(* Logix 5000 project; controller FV vendor 1 type 14 code 217 rev 31.11; software revision 31.00; part 51 of 63 *)
(* tags used below, declared in another part *)
   CWD : CHECKWORD_FLAGS;
   FV_AV1 : PlantItem;   // AV1
   FV_B32 : INT[255];   // PITCH_FLGS YSV pitching control flags
   FV_B32_0_2_OutputBit : BOOL;
   fv_data_file_value_to_move : DINT;
   FV_N12 : INT[255];   // SYS_PARMS System Parameter Fil e
   FV_N141 : INT[255];   // YSV1 DATA
   FV_N142 : INT[255];   // YSV2 DATA
   FV_N143 : INT[255];   // YSV3 DATA
   FV_N30 : INT[255];   // PITCH<PC YSV Pitching data fr om PC
   FV_N31 : INT[255];   // PITCH>PC YSV Pitching data at o PC and control reg isters
   FV_N34 : INT[255];   // PITCH_SV YSV pitching data sa ve file to PC
   FV_N50 : INT[255];   // WASTE<PC
   FV_T33 : TIMER[10];
   FV_YSV1_WTX01_AI : PlantItem;   // YSV1_WTX01
   FV_YSV2_WTX01_AI : PlantItem;   // YSV2_WTX01
   FV_YSV2O : PlantItem;   // YSV2O
   FV_YSV3_WTX01_AI : PlantItem;   // YSV3_WTX01
   FV_YSV3O : PlantItem;   // YSV3O
   FV_YSVPitching_AmountAtEnd : REAL;
   Pitching_transaction_log_delay : DINT;
(* FV_Common, continued *)

ROUTINE FV_PITCH_CP_16   (* ladder *)
   // Reset command interpreter step counter
   0: XIC(S:FS)CLR(FV_N31[16]);
   // RESET
   1: EQU(FV_N31[16],0)MCR();
   2: OTU(FV_B32[0].0);
   3: OTU(FV_B32[0].1);
   4: OTU(FV_B32[0].8);
   5: FLL(0,FV_N31[0],16);
   // Set PCparameter buffer to 'Null' value
   6: FLL(-32768,FV_N30[1],7);
   7: CLR(FV_N30[0]);
   8: MOV(1,FV_N31[16]);
   9: MCR();
   // ALLOW STARTUP DIALOG
   10: EQU(FV_N31[16],1)MCR();
   // Set process status = ready
   11: MOV(1,FV_N31[0]);
   // Allow startup if any vessel is inactive or on storage control only
   12: [[EQU(FV_N141[0],0) ,EQU(FV_N141[0],5) ] ,[EQU(FV_N142[0],0) ,EQU(FV_N142[0],5) ] ,[EQU(FV_N143[0],0) ,EQU(FV_N143[0],5) ] ]OTE(FV_N31[2].0);
   // Advance step if start selected
   13: XIC(FV_N31[2].0)XIC(FV_N30[0].0)MOV(2,FV_N31[16]);
   14: MCR();
   // WAIT FOR STARTUP DIALOG COMPLETE
   15: EQU(FV_N31[16],2)MCR();
   // If YSV1 requested and YSV1 not involved in any other startup dialog set lock flag
   16: EQU(FV_N30[1],1)[EQU(FV_N141[0],0) ,EQU(FV_N141[0],5) ][EQU(FV_N141[4],0) ,XIC(FV_N141[4].2) ]OTE(FV_N141[4].2);
   // If YSV2 requested and YSV2 not involved in any other startup dialog set lock flag
   17: EQU(FV_N30[1],2)[EQU(FV_N142[0],0) ,EQU(FV_N142[0],5) ][EQU(FV_N142[4],0) ,XIC(FV_N142[4].2) ]OTE(FV_N142[4].2);
   // If YSV3 requested and YSV3 not involved in any other startup dialog set lock flag
   18: EQU(FV_N30[1],3)[EQU(FV_N143[0],0) ,EQU(FV_N143[0],5) ][EQU(FV_N143[4],0) ,XIC(FV_N143[4].2) ]OTE(FV_N143[4].2);
   // Allow start confirmed button if selected YSV could be locked
   19: [XIC(FV_N141[4].2) ,XIC(FV_N142[4].2) ,XIC(FV_N143[4].2) ]OTE(FV_N31[2].1);
   // Startup dialog guard timer
   20: TON(FV_T33[0],?,?);
   // Reset command processor if dialog cancel selected or startup dialog timer expired
   21: [XIC(FV_N30[0].15) ,XIC(FV_T33[0].DN) ]CLR(FV_N31[16]);
   // Advance step if start available and selected
   22: XIC(FV_N30[0].1)XIC(FV_N31[2].1)[MOV(3,FV_N31[16]) ,CLR(FV_N30[0]) ];
   23: MCR();
   // COMPLETE STARTUP DIALOG
   24: EQU(FV_N31[16],3)MCR();
   // If YSV 1 selected, save YSV1 status
   25: EQU(FV_N30[1],1)MOV(FV_N141[0],FV_N31[12]);
   // If YSV2 selected, save YSV2 status
   26: EQU(FV_N50[1],2)MOV(FV_N142[0],FV_N31[12]);
   // If YSV 3 selected, save YSV3 status
   27: EQU(FV_N50[1],3)MOV(FV_N143[0],FV_N31[12]);
   // If YSV 1 selected, set YSV1 status = Pitching
   28: EQU(FV_N30[1],1)MOV(2,FV_N141[0]);
   // If YSV 2 selected, set YSV2 status = Pitching
   29: EQU(FV_N30[1],2)MOV(2,FV_N142[0]);
   // If YSV 3 selected, set YSV3 status = Pitching
   30: EQU(FV_N30[1],3)MOV(2,FV_N143[0]);
   // Set YSV Pitching Process Status = Running
   31: MOV(2,FV_N31[0]);
   32: OTL(FV_B32[0].0);
   33: OTL(FV_B32[0].1);
   34: OTL(FV_N31[2].2);
   35: MOV(10,FV_N31[1]);
   36: MOV(10,FV_N31[3]);
   37: MOV(-1,FV_N31[16]);
   38: CLR(FV_N30[0]);
   39: MCR();
   // HANDLE STOP BUTTON
   40: XIC(FV_N30[0].2)XIC(FV_N31[2].2)MCR();
   41: OTU(FV_B32[0].1);
   42: OTU(FV_N31[2].2);
   43: OTL(FV_N31[2].3);
   44: OTL(FV_N31[2].4);
   45: MOV(3,FV_N31[0]);
   46: MOV(0,FV_N31[1]);
   47: CLR(FV_N30[0]);
   48: MCR();
   // HANDLE CONTINUE BUTTON
   49: XIC(FV_N30[0].3)XIC(FV_N31[2].3)MCR();
   50: OTL(FV_B32[0].1);
   51: OTL(FV_N31[2].2);
   52: OTU(FV_N31[2].3);
   // Reset process alarm and parameters
   53: OTU(FV_N31[2].4);
   54: FLL(0,FV_N31[4],4);
   55: MOV(2,FV_N31[0]);
   // Set current Step = Restart Step
   56: MOV(FV_N31[3],FV_N31[1]);
   57: CLR(FV_N30[0]);
   58: MCR();
   // HANDLE ABORT BUTTON
   59: XIC(FV_N30[0].4)XIC(FV_N31[2].4)MCR();
   60: OTU(FV_B32[0].0);
   // Set rouser control mode for current vessel to automatic
   61: JSR(FV_Set_FV_Datafile_Value,3,0,FV_N31[15],3);
   // If FV attemporation control is waiting, set it to rise phase
   62: JSR(FV_Get_FV_Datafile_Value,2,FV_N31[13],24)EQU(fv_data_file_value_to_move,8)JSR(FV_Set_FV_Datafile_Value,3,1,FV_N31[13],24);
   // Set YSV's operation to status prior to pitching
   63: JSR(FV_Set_FV_Datafile_Value,3,FV_N31[12],FV_N31[15],0);
   64: CLR(FV_N31[16]);
   65: CLR(FV_N30[0]);
   66: MCR();
   // Copy step number for PC to display if running
   67: XIC(FV_B32[0].1)MOV(FV_N31[1],FV_N31[9]);
END_ROUTINE

ROUTINE FV_PITCH_MC_15   (* ladder *)
   // Run Pitching command interpreter
   0: JSR(FV_PITCH_CP_16,0);
   // Run Pitching Process If Active
   1: XIC(FV_B32[0].0)JSR(FV_PITCH_PRO_17,0);
   // PostScan Pitching Process If not active
   2: XIO(FV_B32[0].0)OSR(FV_B32[0].2,FV_B32_0_2_OutputBit)XIC(FV_B32_0_2_OutputBit)JSR(FV_PITCH_PRO_17,0);
END_ROUTINE

ROUTINE FV_PITCH_PRO_17   (* ladder *)
   // YSV PITCHING - STEP 10 - Initialize
   0: XIC(FV_B32[0].1)EQU(FV_N31[1],10)MCR();
   // Set restart step for this process
   1: MOV(10,FV_N31[3]);
   // Make pointer to selected YSV's data file
   2: ADD(FV_N30[1],140,FV_N31[15]);
   // Make pointer to YSV's Attemporation Data File
   3: ADD(FV_N30[1],135,FV_N31[14]);
   // Make pointer to FV's attemporation data file
   4: [ADD(FV_N30[3],110,FV_N31[13]) ,LIM(226,FV_N30[3],231) SUB(FV_N30[3],80,FV_N31[13]) ];
   // Save YSV volume at start of transfer
   5: JSR(FV_Get_FV_Datafile_Value,2,FV_N31[15],5)MOV(fv_data_file_value_to_move,FV_N31[17]);
   // Calculate maximum allowed volume in YSV before alarm
   6: ADD(FV_N31[17],FV_N12[4],FV_N31[18]);
   // Calculate volume at which to stop pitching. If < 0 , set to zero
   7: [SUB(FV_N31[17],FV_N30[2],FV_N31[21]) ,LES(FV_N31[21],0) MOV(0,FV_N31[21]) ];
   // Advance to next step
   8: MOV(20,FV_N31[1]);
   9: MCR();
   // Request inlet / outlet valve on correct vessel
   10: [EQU(FV_N30[1],1) MOV(FV_YSV1_WTX01_AI.Scaled,FV_YSVPitching_AmountAtEnd) ,EQU(FV_N30[1],2) MOV(FV_YSV2_WTX01_AI.Scaled,FV_YSVPitching_AmountAtEnd) ,EQU(FV_N30[1],3) MOV(FV_YSV3_WTX01_AI.Scaled,FV_YSVPitching_AmountAtEnd) ];
   // YSV PITCHING - STEP 20 - Pitch to FV
   11: XIC(FV_B32[0].1)EQU(FV_N31[1],20)MCR();
   // Set restart step for this process
   12: MOV(20,FV_N31[3]);
   // Request inlet / outlet valve on correct vessel
   13: [EQU(FV_N30[1],1) OTE(FV_AV1.DriveBits.2) ,EQU(FV_N30[1],2) OTE(FV_YSV2O.DriveBits.2) ,EQU(FV_N30[1],3) OTE(FV_YSV3O.DriveBits.2) ];
   // Generate alarm if YSV weight increases whilst vessel is transfering
   14: JSR(FV_Get_FV_Datafile_Value,2,FV_N31[15],5)GRT(fv_data_file_value_to_move,FV_N31[18])[MOV(200,FV_N31[4]) ,MOV(FV_N30[1],FV_N31[5]) ];
   // Check for low pitching rate if vessel > low level value
   15: JSR(FV_Get_FV_Datafile_Value,2,FV_N31[15],5)GRT(fv_data_file_value_to_move,100)XIO(FV_T33[1].DN)[TON(FV_T33[1],?,?) ,EQU(FV_T33[1].ACC,0) JSR(FV_Get_FV_Datafile_Value,2,FV_N31[15],5) MOV(fv_data_file_value_to_move,FV_N31[19]) ,XIC(FV_T33[1].DN) [JSR(FV_Get_FV_Datafile_Value,2,FV_N31[15],5) SUB(FV_N31[19],fv_data_file_value_to_move,FV_N31[20]) ,LES(FV_N31[20],FV_N12[5]) [MOV(201,FV_N31[4]) ,MOV(FV_N30[1],FV_N31[5]) ] ] ];
   // Calculate  volume pitched so far for SCADA display
   16: JSR(FV_Get_FV_Datafile_Value,2,FV_N31[15],5)SUB(FV_N31[17],fv_data_file_value_to_move,FV_N31[10]);
   // Advance to next step if target volume pitched
   17: LEQ(fv_data_file_value_to_move,FV_N31[21])MOV(30,FV_N31[1]);
   // Allow operator to select process end button
   18: OTE(FV_N31[2].5);
   // Advance to next step when End selected
   19: XIC(FV_N30[0].5)MOV(30,FV_N31[1]);
   20: MCR();
   // YSV PITCHING - STEP 30 - Save Pitched Volume
   21: XIC(FV_B32[0].1)EQU(FV_N31[1],30)MCR();
   // Delay to allow vessel outlet to close and  weight to steady
   22: TON(FV_T33[2],?,?);
   // Calculate and Save volume pitched
   23: XIC(FV_T33[2].DN)JSR(FV_Get_FV_Datafile_Value,2,FV_N31[15],5)SUB(FV_N31[17],fv_data_file_value_to_move,FV_N34[2]);
   24: XIC(FV_T33[2].DN)MOV(40,FV_N31[1]);
   25: MCR();
   // YSV PITCHING - STEP 40 - Reset YSV and FV
   26: XIC(FV_B32[0].1)EQU(FV_N31[1],40)MCR();
   // Set rouser control mode for current vessel to automatic
   27: JSR(FV_Set_FV_Datafile_Value,3,0,FV_N31[15],3);
   // Set YSV status to storage operation
   28: JSR(FV_Set_FV_Datafile_Value,3,5,FV_N31[15],0);
   // If FV attemporation control is waiting, set it to rise phase
   29: JSR(FV_Get_FV_Datafile_Value,2,FV_N31[13],24)EQU(fv_data_file_value_to_move,8)JSR(FV_Set_FV_Datafile_Value,3,1,FV_N31[13],24);
   30: MOV(50,FV_N31[1]);
   31: MCR();
   // YSV PITCHING - STEP 50 - Save Data
   32: XIC(FV_B32[0].1)EQU(FV_N31[1],50)MCR();
   // Save YSV number which pitched to PC
   33: MOV(FV_N30[1],FV_N34[1]);
   // Save FV number which was pitched to PC
   34: MOV(FV_N30[3],FV_N34[3]);
   // Set Save data flag to PC
   35: MOV(1,FV_N34[0]);
   36: MOV(1,Pitching_transaction_log_delay);
   37: CLR(FV_N31[16]);
   38: MCR();
   // CHECK FOR ALARM CONDITIONS
   39: XIC(FV_B32[0].1)MCR();
   40: EQU(FV_N30[1],1)XIC(FV_AV1.CW.[CWD.FAULT])OTU(FV_B32[0].1);
   41: GRT(FV_N31[4],0)OTU(FV_B32[0].1);
   42: XIO(FV_B32[0].1)[MOV(4,FV_N31[0]) ,OTU(FV_N31[2].2) ,OTL(FV_N31[2].3) ,OTL(FV_N31[2].4) ,MOV(0,FV_N31[1]) ];
   43: MCR();
END_ROUTINE
